TYPE "From Excel: Data"
VERSION : 0.1
   STRUCT
      kp8Stns : Array[0.."kp8StnCount"] of "From Excel: Codes Single Wip";
      hmiStns : Array[0.."hmi_station_count"] of "From Excel: Codes Multiple Wips";
   END_STRUCT;
   // hmiStns[0].wip[40].pnCode[3] := 1000;
   // hmiStns[0].wip[0].pnCode[2] := 20000;
   // hmiStns[0].wip[0].pnCode[1] := 244000;
   // hmiStns[0].wip[0].pnCode[0] := 1000;
   // hmiStns[0].pStn := 25;
   // kp8Stns[0].pStn := 0;
   // kp8Stns[0].pnCode[7] := 169000;
   // kp8Stns[2].pStn := 2;
   // kp8Stns[3].pStn := 3;
   // kp8Stns[4].pStn := 4;
   // kp8Stns[5].pStn := 5;
   // kp8Stns[7].pStn := 7;
   // kp8Stns[8].pStn := 8;
   // kp8Stns[9].pStn := 9;
   // kp8Stns[10].pStn := 10;
   // kp8Stns[11].pStn := 11;
   // kp8Stns[12].pStn := 12;
   // kp8Stns[13].pStn := 13;
   // kp8Stns[14].pStn := 14;
   // kp8Stns[15].pStn := 15;
   // kp8Stns[16].pStn := 16;
   // kp8Stns[17].pStn := 17;
   // kp8Stns[18].pStn := 18;
   // kp8Stns[19].pStn := 19;
   // kp8Stns[20].pStn := 20;
   // kp8Stns[21].pStn := 21;
   // kp8Stns[22].pStn := 22;
   // kp8Stns[23].pStn := 23;
   // kp8Stns[24].pStn := 24;
   // kp8Stns[6].pStn := 6;
   // kp8Stns[25].pStn := 30;
   // kp8Stns[26].pStn := 31;
   // kp8Stns[27].pStn := 32;
   // kp8Stns[28].pStn := 33;
   // kp8Stns[30].pStn := 35;
   // kp8Stns[31].pStn := 36;
   // kp8Stns[32].pStn := 37;
   // kp8Stns[29].pStn := 34;
   // kp8Stns[33].pStn := 38;
   // hmiStns[0].wip[40].pnCode[2] := 1000;
   // hmiStns[0].wip[40].pnCode[1] := 1000;
   // hmiStns[0].wip[40].pnCode[0] := 1000;
   // hmiStns[0].wip[39].pnCode[7] := 1000;
   // hmiStns[0].wip[39].pnCode[6] := 1000;
   // hmiStns[0].wip[39].pnCode[5] := 1000;
   // hmiStns[0].wip[39].pnCode[4] := 1000;
   // hmiStns[0].wip[39].pnCode[3] := 1000;
   // hmiStns[0].wip[39].pnCode[2] := 1000;
   // hmiStns[0].wip[39].pnCode[1] := 1000;
   // hmiStns[0].wip[39].pnCode[0] := 1000;
   // hmiStns[0].wip[38].pnCode[7] := 1000;
   // hmiStns[0].wip[38].pnCode[6] := 1000;
   // hmiStns[0].wip[38].pnCode[5] := 1000;
   // hmiStns[0].wip[38].pnCode[4] := 1000;
   // hmiStns[0].wip[38].pnCode[3] := 1000;
   // hmiStns[0].wip[38].pnCode[2] := 1000;
   // hmiStns[0].wip[38].pnCode[1] := 1000;
   // hmiStns[0].wip[38].pnCode[0] := 1000;
   // hmiStns[0].wip[37].pnCode[7] := 1000;
   // hmiStns[0].wip[37].pnCode[6] := 1000;
   // hmiStns[0].wip[37].pnCode[5] := 1000;
   // hmiStns[0].wip[37].pnCode[4] := 1000;
   // hmiStns[0].wip[37].pnCode[3] := 1000;
   // hmiStns[0].wip[37].pnCode[2] := 1000;
   // hmiStns[0].wip[37].pnCode[1] := 1000;
   // hmiStns[0].wip[37].pnCode[0] := 1000;
   // hmiStns[0].wip[36].pnCode[7] := 1000;
   // hmiStns[0].wip[36].pnCode[6] := 1000;
   // hmiStns[0].wip[36].pnCode[5] := 1000;
   // hmiStns[0].wip[36].pnCode[4] := 1000;
   // hmiStns[0].wip[36].pnCode[3] := 1000;
   // hmiStns[0].wip[36].pnCode[2] := 1000;
   // hmiStns[0].wip[36].pnCode[1] := 1000;
   // hmiStns[0].wip[36].pnCode[0] := 1000;
   // hmiStns[0].wip[35].pnCode[7] := 1000;
   // hmiStns[0].wip[35].pnCode[6] := 1000;
   // hmiStns[0].wip[35].pnCode[5] := 1000;
   // hmiStns[0].wip[35].pnCode[4] := 1000;
   // hmiStns[0].wip[35].pnCode[3] := 1000;
   // hmiStns[0].wip[35].pnCode[2] := 1000;
   // hmiStns[0].wip[35].pnCode[1] := 1000;
   // hmiStns[0].wip[35].pnCode[0] := 1000;
   // hmiStns[0].wip[34].pnCode[7] := 1000;
   // hmiStns[0].wip[34].pnCode[6] := 1000;
   // hmiStns[0].wip[34].pnCode[5] := 1000;
   // hmiStns[0].wip[34].pnCode[4] := 1000;
   // hmiStns[0].wip[34].pnCode[3] := 1000;
   // hmiStns[0].wip[34].pnCode[2] := 1000;
   // hmiStns[0].wip[34].pnCode[1] := 1000;
   // hmiStns[0].wip[34].pnCode[0] := 1000;
   // hmiStns[0].wip[33].pnCode[7] := 1000;
   // hmiStns[0].wip[33].pnCode[6] := 1000;
   // hmiStns[0].wip[33].pnCode[5] := 1000;
   // hmiStns[0].wip[33].pnCode[4] := 1000;
   // hmiStns[0].wip[33].pnCode[3] := 1000;
   // hmiStns[0].wip[33].pnCode[2] := 1000;
   // hmiStns[0].wip[33].pnCode[1] := 1000;
   // hmiStns[0].wip[33].pnCode[0] := 1000;
   // hmiStns[0].wip[32].pnCode[7] := 1000;
   // hmiStns[0].wip[32].pnCode[6] := 1000;
   // hmiStns[0].wip[32].pnCode[5] := 1000;
   // hmiStns[0].wip[32].pnCode[4] := 1000;
   // hmiStns[0].wip[32].pnCode[3] := 1000;
   // hmiStns[0].wip[32].pnCode[2] := 1000;
   // hmiStns[0].wip[32].pnCode[1] := 1000;
   // hmiStns[0].wip[32].pnCode[0] := 1000;
   // hmiStns[0].wip[31].pnCode[7] := 1000;
   // hmiStns[0].wip[31].pnCode[6] := 1000;
   // hmiStns[0].wip[31].pnCode[5] := 1000;
   // hmiStns[0].wip[31].pnCode[4] := 1000;
   // hmiStns[0].wip[31].pnCode[3] := 1000;
   // hmiStns[0].wip[31].pnCode[2] := 1000;
   // hmiStns[0].wip[31].pnCode[1] := 1000;
   // hmiStns[0].wip[31].pnCode[0] := 1000;
   // hmiStns[0].wip[30].pnCode[7] := 1000;
   // hmiStns[0].wip[30].pnCode[6] := 1000;
   // hmiStns[0].wip[30].pnCode[5] := 1000;
   // hmiStns[0].wip[30].pnCode[4] := 1000;
   // hmiStns[0].wip[30].pnCode[3] := 1000;
   // hmiStns[0].wip[30].pnCode[2] := 1000;
   // hmiStns[0].wip[30].pnCode[1] := 1000;
   // hmiStns[0].wip[30].pnCode[0] := 1000;
   // hmiStns[0].wip[29].pnCode[7] := 1000;
   // hmiStns[0].wip[29].pnCode[6] := 1000;
   // hmiStns[0].wip[29].pnCode[5] := 1000;
   // hmiStns[0].wip[29].pnCode[4] := 1000;
   // hmiStns[0].wip[29].pnCode[3] := 1000;
   // hmiStns[0].wip[29].pnCode[2] := 1000;
   // hmiStns[0].wip[29].pnCode[1] := 1000;
   // hmiStns[0].wip[29].pnCode[0] := 1000;
   // hmiStns[0].wip[28].pnCode[7] := 1000;
   // hmiStns[0].wip[28].pnCode[6] := 1000;
   // hmiStns[0].wip[28].pnCode[5] := 1000;
   // hmiStns[0].wip[28].pnCode[4] := 1000;
   // hmiStns[0].wip[28].pnCode[3] := 1000;
   // hmiStns[0].wip[28].pnCode[2] := 1000;
   // hmiStns[0].wip[28].pnCode[1] := 1000;
   // hmiStns[0].wip[28].pnCode[0] := 1000;
   // hmiStns[0].wip[27].pnCode[7] := 1000;
   // hmiStns[0].wip[27].pnCode[6] := 1000;
   // hmiStns[0].wip[27].pnCode[5] := 1000;
   // hmiStns[0].wip[27].pnCode[4] := 1000;
   // hmiStns[0].wip[27].pnCode[3] := 1000;
   // hmiStns[0].wip[27].pnCode[2] := 1000;
   // hmiStns[0].wip[27].pnCode[1] := 1000;
   // hmiStns[0].wip[27].pnCode[0] := 1000;
   // hmiStns[0].wip[26].pnCode[7] := 1000;
   // hmiStns[0].wip[26].pnCode[6] := 1000;
   // hmiStns[0].wip[26].pnCode[5] := 1000;
   // hmiStns[0].wip[26].pnCode[4] := 1000;
   // hmiStns[0].wip[26].pnCode[3] := 1000;
   // hmiStns[0].wip[26].pnCode[2] := 1000;
   // hmiStns[0].wip[26].pnCode[1] := 1000;
   // hmiStns[0].wip[26].pnCode[0] := 1000;
   // hmiStns[0].wip[25].pnCode[7] := 1000;
   // hmiStns[0].wip[25].pnCode[6] := 1000;
   // hmiStns[0].wip[25].pnCode[5] := 1000;
   // hmiStns[0].wip[25].pnCode[4] := 1000;
   // hmiStns[0].wip[25].pnCode[3] := 1000;
   // hmiStns[0].wip[25].pnCode[2] := 1000;
   // hmiStns[0].wip[25].pnCode[1] := 1000;
   // hmiStns[0].wip[25].pnCode[0] := 1000;
   // hmiStns[0].wip[24].pnCode[7] := 1000;
   // hmiStns[0].wip[24].pnCode[6] := 1000;
   // hmiStns[0].wip[24].pnCode[5] := 1000;
   // hmiStns[0].wip[24].pnCode[4] := 1000;
   // hmiStns[0].wip[24].pnCode[3] := 1000;
   // hmiStns[0].wip[24].pnCode[2] := 1000;
   // hmiStns[0].wip[24].pnCode[1] := 1000;
   // hmiStns[0].wip[24].pnCode[0] := 1000;
   // hmiStns[0].wip[23].pnCode[7] := 223000;
   // hmiStns[0].wip[23].pnCode[6] := 220000;
   // hmiStns[0].wip[23].pnCode[5] := 1000;
   // hmiStns[0].wip[23].pnCode[4] := 1000;
   // hmiStns[0].wip[23].pnCode[3] := 1000;
   // hmiStns[0].wip[23].pnCode[2] := 221000;
   // hmiStns[0].wip[23].pnCode[1] := 244000;
   // hmiStns[0].wip[23].pnCode[0] := 1000;
   // hmiStns[0].wip[22].pnCode[7] := 223000;
   // hmiStns[0].wip[22].pnCode[6] := 222000;
   // hmiStns[0].wip[22].pnCode[5] := 1000;
   // hmiStns[0].wip[22].pnCode[4] := 1000;
   // hmiStns[0].wip[22].pnCode[3] := 220000;
   // hmiStns[0].wip[22].pnCode[2] := 1000;
   // hmiStns[0].wip[22].pnCode[1] := 244000;
   // hmiStns[0].wip[22].pnCode[0] := 1000;
   // hmiStns[0].wip[21].pnCode[7] := 31000;
   // hmiStns[0].wip[21].pnCode[6] := 51000;
   // hmiStns[0].wip[21].pnCode[5] := 1000;
   // hmiStns[0].wip[21].pnCode[4] := 1000;
   // hmiStns[0].wip[21].pnCode[3] := 32000;
   // hmiStns[0].wip[21].pnCode[2] := 1000;
   // hmiStns[0].wip[21].pnCode[1] := 244000;
   // hmiStns[0].wip[21].pnCode[0] := 1000;
   // hmiStns[0].wip[20].pnCode[7] := 17000;
   // hmiStns[0].wip[20].pnCode[6] := 25000;
   // hmiStns[0].wip[20].pnCode[5] := 1000;
   // hmiStns[0].wip[20].pnCode[4] := 1000;
   // hmiStns[0].wip[20].pnCode[3] := 1000;
   // hmiStns[0].wip[20].pnCode[2] := 18000;
   // hmiStns[0].wip[20].pnCode[1] := 244000;
   // hmiStns[0].wip[20].pnCode[0] := 1000;
   // hmiStns[0].wip[19].pnCode[7] := 227000;
   // hmiStns[0].wip[19].pnCode[6] := 226000;
   // hmiStns[0].wip[19].pnCode[5] := 1000;
   // hmiStns[0].wip[19].pnCode[4] := 1000;
   // hmiStns[0].wip[19].pnCode[3] := 1000;
   // hmiStns[0].wip[19].pnCode[2] := 225000;
   // hmiStns[0].wip[19].pnCode[1] := 244000;
   // hmiStns[0].wip[19].pnCode[0] := 1000;
   // hmiStns[0].wip[18].pnCode[7] := 224000;
   // hmiStns[0].wip[18].pnCode[6] := 219000;
   // hmiStns[0].wip[18].pnCode[5] := 1000;
   // hmiStns[0].wip[18].pnCode[4] := 1000;
   // hmiStns[0].wip[18].pnCode[3] := 1000;
   // hmiStns[0].wip[18].pnCode[2] := 199000;
   // hmiStns[0].wip[18].pnCode[1] := 244000;
   // hmiStns[0].wip[18].pnCode[0] := 1000;
   // hmiStns[0].wip[17].pnCode[7] := 223000;
   // hmiStns[0].wip[17].pnCode[6] := 220000;
   // hmiStns[0].wip[17].pnCode[5] := 1000;
   // hmiStns[0].wip[17].pnCode[4] := 1000;
   // hmiStns[0].wip[17].pnCode[3] := 1000;
   // hmiStns[0].wip[17].pnCode[2] := 198000;
   // hmiStns[0].wip[17].pnCode[1] := 244000;
   // hmiStns[0].wip[17].pnCode[0] := 1000;
   // hmiStns[0].wip[16].pnCode[7] := 224000;
   // hmiStns[0].wip[16].pnCode[6] := 219000;
   // hmiStns[0].wip[16].pnCode[5] := 1000;
   // hmiStns[0].wip[16].pnCode[4] := 1000;
   // hmiStns[0].wip[16].pnCode[3] := 1000;
   // hmiStns[0].wip[16].pnCode[2] := 218000;
   // hmiStns[0].wip[16].pnCode[1] := 244000;
   // hmiStns[0].wip[16].pnCode[0] := 1000;
   // hmiStns[0].wip[15].pnCode[7] := 37000;
   // hmiStns[0].wip[15].pnCode[6] := 36000;
   // hmiStns[0].wip[15].pnCode[5] := 1000;
   // hmiStns[0].wip[15].pnCode[4] := 1000;
   // hmiStns[0].wip[15].pnCode[3] := 1000;
   // hmiStns[0].wip[15].pnCode[2] := 100000;
   // hmiStns[0].wip[15].pnCode[1] := 244000;
   // hmiStns[0].wip[15].pnCode[0] := 1000;
   // hmiStns[0].wip[14].pnCode[7] := 37000;
   // hmiStns[0].wip[14].pnCode[6] := 43000;
   // hmiStns[0].wip[14].pnCode[5] := 1000;
   // hmiStns[0].wip[14].pnCode[4] := 1000;
   // hmiStns[0].wip[14].pnCode[3] := 1000;
   // hmiStns[0].wip[14].pnCode[2] := 100000;
   // hmiStns[0].wip[14].pnCode[1] := 244000;
   // hmiStns[0].wip[14].pnCode[0] := 1000;
   // hmiStns[0].wip[13].pnCode[7] := 45000;
   // hmiStns[0].wip[13].pnCode[6] := 39000;
   // hmiStns[0].wip[13].pnCode[5] := 1000;
   // hmiStns[0].wip[13].pnCode[4] := 1000;
   // hmiStns[0].wip[13].pnCode[3] := 1000;
   // hmiStns[0].wip[13].pnCode[2] := 99000;
   // hmiStns[0].wip[13].pnCode[1] := 244000;
   // hmiStns[0].wip[13].pnCode[0] := 1000;
   // hmiStns[0].wip[12].pnCode[7] := 72000;
   // hmiStns[0].wip[12].pnCode[6] := 32000;
   // hmiStns[0].wip[12].pnCode[5] := 1000;
   // hmiStns[0].wip[12].pnCode[4] := 1000;
   // hmiStns[0].wip[12].pnCode[3] := 1000;
   // hmiStns[0].wip[12].pnCode[2] := 85000;
   // hmiStns[0].wip[12].pnCode[1] := 244000;
   // hmiStns[0].wip[12].pnCode[0] := 1000;
   // hmiStns[0].wip[11].pnCode[7] := 19000;
   // hmiStns[0].wip[11].pnCode[6] := 26000;
   // hmiStns[0].wip[11].pnCode[5] := 1000;
   // hmiStns[0].wip[11].pnCode[4] := 1000;
   // hmiStns[0].wip[11].pnCode[3] := 1000;
   // hmiStns[0].wip[11].pnCode[2] := 58000;
   // hmiStns[0].wip[11].pnCode[1] := 244000;
   // hmiStns[0].wip[11].pnCode[0] := 1000;
   // hmiStns[0].wip[10].pnCode[7] := 72000;
   // hmiStns[0].wip[10].pnCode[6] := 32000;
   // hmiStns[0].wip[10].pnCode[5] := 1000;
   // hmiStns[0].wip[10].pnCode[4] := 1000;
   // hmiStns[0].wip[10].pnCode[3] := 1000;
   // hmiStns[0].wip[10].pnCode[2] := 54000;
   // hmiStns[0].wip[10].pnCode[1] := 244000;
   // hmiStns[0].wip[10].pnCode[0] := 1000;
   // hmiStns[0].wip[9].pnCode[7] := 74000;
   // hmiStns[0].wip[9].pnCode[6] := 32000;
   // hmiStns[0].wip[9].pnCode[5] := 1000;
   // hmiStns[0].wip[9].pnCode[4] := 1000;
   // hmiStns[0].wip[9].pnCode[3] := 1000;
   // hmiStns[0].wip[9].pnCode[2] := 53000;
   // hmiStns[0].wip[9].pnCode[1] := 244000;
   // hmiStns[0].wip[9].pnCode[0] := 1000;
   // hmiStns[0].wip[8].pnCode[7] := 19000;
   // hmiStns[0].wip[8].pnCode[6] := 26000;
   // hmiStns[0].wip[8].pnCode[5] := 1000;
   // hmiStns[0].wip[8].pnCode[4] := 1000;
   // hmiStns[0].wip[8].pnCode[3] := 1000;
   // hmiStns[0].wip[8].pnCode[2] := 52000;
   // hmiStns[0].wip[8].pnCode[1] := 244000;
   // hmiStns[0].wip[8].pnCode[0] := 1000;
   // hmiStns[0].wip[7].pnCode[7] := 45000;
   // hmiStns[0].wip[7].pnCode[6] := 39000;
   // hmiStns[0].wip[7].pnCode[5] := 1000;
   // hmiStns[0].wip[7].pnCode[4] := 1000;
   // hmiStns[0].wip[7].pnCode[3] := 1000;
   // hmiStns[0].wip[7].pnCode[2] := 44000;
   // hmiStns[0].wip[7].pnCode[1] := 244000;
   // hmiStns[0].wip[7].pnCode[0] := 1000;
   // hmiStns[0].wip[6].pnCode[7] := 37000;
   // hmiStns[0].wip[6].pnCode[6] := 43000;
   // hmiStns[0].wip[6].pnCode[5] := 1000;
   // hmiStns[0].wip[6].pnCode[4] := 1000;
   // hmiStns[0].wip[6].pnCode[3] := 1000;
   // hmiStns[0].wip[6].pnCode[2] := 46000;
   // hmiStns[0].wip[6].pnCode[1] := 244000;
   // hmiStns[0].wip[6].pnCode[0] := 1000;
   // hmiStns[0].wip[5].pnCode[7] := 37000;
   // hmiStns[0].wip[5].pnCode[6] := 43000;
   // hmiStns[0].wip[5].pnCode[5] := 1000;
   // hmiStns[0].wip[5].pnCode[4] := 1000;
   // hmiStns[0].wip[5].pnCode[3] := 1000;
   // hmiStns[0].wip[5].pnCode[2] := 38000;
   // hmiStns[0].wip[5].pnCode[1] := 244000;
   // hmiStns[0].wip[5].pnCode[0] := 1000;
   // hmiStns[0].wip[4].pnCode[7] := 37000;
   // hmiStns[0].wip[4].pnCode[6] := 36000;
   // hmiStns[0].wip[4].pnCode[5] := 1000;
   // hmiStns[0].wip[4].pnCode[4] := 1000;
   // hmiStns[0].wip[4].pnCode[3] := 1000;
   // hmiStns[0].wip[4].pnCode[2] := 46000;
   // hmiStns[0].wip[4].pnCode[1] := 244000;
   // hmiStns[0].wip[4].pnCode[0] := 1000;
   // hmiStns[0].wip[3].pnCode[7] := 33000;
   // hmiStns[0].wip[3].pnCode[6] := 42000;
   // hmiStns[0].wip[3].pnCode[5] := 15000;
   // hmiStns[0].wip[3].pnCode[4] := 1000;
   // hmiStns[0].wip[3].pnCode[3] := 14000;
   // hmiStns[0].wip[3].pnCode[2] := 48000;
   // hmiStns[0].wip[3].pnCode[1] := 244000;
   // hmiStns[0].wip[3].pnCode[0] := 1000;
   // hmiStns[0].wip[2].pnCode[7] := 40000;
   // hmiStns[0].wip[2].pnCode[6] := 39000;
   // hmiStns[0].wip[2].pnCode[5] := 1000;
   // hmiStns[0].wip[2].pnCode[4] := 1000;
   // hmiStns[0].wip[2].pnCode[3] := 1000;
   // hmiStns[0].wip[2].pnCode[2] := 41000;
   // hmiStns[0].wip[2].pnCode[1] := 244000;
   // hmiStns[0].wip[2].pnCode[0] := 1000;
   // hmiStns[0].wip[1].pnCode[7] := 37000;
   // hmiStns[0].wip[1].pnCode[6] := 36000;
   // hmiStns[0].wip[1].pnCode[5] := 1000;
   // hmiStns[0].wip[1].pnCode[4] := 1000;
   // hmiStns[0].wip[1].pnCode[3] := 1000;
   // hmiStns[0].wip[1].pnCode[2] := 38000;
   // hmiStns[0].wip[1].pnCode[1] := 244000;
   // hmiStns[0].wip[1].pnCode[0] := 1000;
   // hmiStns[0].wip[0].pnCode[7] := 19000;
   // hmiStns[0].wip[0].pnCode[6] := 26000;
   // hmiStns[0].wip[0].pnCode[5] := 1000;
   // hmiStns[0].wip[0].pnCode[4] := 1000;
   // hmiStns[0].wip[0].pnCode[3] := 1000;
   // kp8Stns[1].pnCode[0] := 1000;
   // kp8Stns[0].pnCode[1] := 1000;
   // kp8Stns[0].pnCode[0] := 1000;
   // kp8Stns[0].pnCode[2] := 1000;
   // kp8Stns[0].pnCode[3] := 173000;
   // kp8Stns[0].pnCode[4] := 1000;
   // kp8Stns[0].pnCode[5] := 1000;
   // kp8Stns[0].pnCode[6] := 1000;
   // kp8Stns[1].pnCode[1] := 1000;
   // kp8Stns[1].pnCode[2] := 184000;
   // kp8Stns[1].pnCode[3] := 210000;
   // kp8Stns[1].pnCode[4] := 1000;
   // kp8Stns[1].pnCode[5] := 1000;
   // kp8Stns[1].pnCode[6] := 181000;
   // kp8Stns[1].pnCode[7] := 167000;
   // kp8Stns[1].pStn := 1;
   // kp8Stns[2].pnCode[0] := 1000;
   // kp8Stns[2].pnCode[1] := 183000;
   // kp8Stns[2].pnCode[2] := 182000;
   // kp8Stns[2].pnCode[3] := 216000;
   // kp8Stns[2].pnCode[4] := 1000;
   // kp8Stns[2].pnCode[5] := 185000;
   // kp8Stns[2].pnCode[6] := 217000;
   // kp8Stns[2].pnCode[7] := 215000;
   // kp8Stns[3].pnCode[0] := 1000;
   // kp8Stns[3].pnCode[1] := 193000;
   // kp8Stns[3].pnCode[2] := 192000;
   // kp8Stns[3].pnCode[3] := 189000;
   // kp8Stns[3].pnCode[4] := 1000;
   // kp8Stns[3].pnCode[5] := 191000;
   // kp8Stns[3].pnCode[6] := 188000;
   // kp8Stns[3].pnCode[7] := 190000;
   // kp8Stns[4].pnCode[0] := 1000;
   // kp8Stns[4].pnCode[1] := 1000;
   // kp8Stns[4].pnCode[2] := 1000;
   // kp8Stns[4].pnCode[3] := 1000;
   // kp8Stns[4].pnCode[4] := 1000;
   // kp8Stns[4].pnCode[5] := 1000;
   // kp8Stns[4].pnCode[6] := 1000;
   // kp8Stns[4].pnCode[7] := 195000;
   // kp8Stns[5].pnCode[0] := 1000;
   // kp8Stns[5].pnCode[1] := 194000;
   // kp8Stns[5].pnCode[2] := 196000;
   // kp8Stns[5].pnCode[3] := 177000;
   // kp8Stns[5].pnCode[4] := 1000;
   // kp8Stns[5].pnCode[5] := 197000;
   // kp8Stns[5].pnCode[6] := 178000;
   // kp8Stns[5].pnCode[7] := 176000;
   // kp8Stns[6].pnCode[0] := 1000;
   // kp8Stns[6].pnCode[1] := 209000;
   // kp8Stns[6].pnCode[2] := 208000;
   // kp8Stns[6].pnCode[3] := 211000;
   // kp8Stns[6].pnCode[4] := 1000;
   // kp8Stns[6].pnCode[5] := 212000;
   // kp8Stns[6].pnCode[6] := 207000;
   // kp8Stns[6].pnCode[7] := 206000;
   // kp8Stns[7].pnCode[0] := 1000;
   // kp8Stns[7].pnCode[1] := 1000;
   // kp8Stns[7].pnCode[2] := 1000;
   // kp8Stns[7].pnCode[3] := 175000;
   // kp8Stns[7].pnCode[4] := 1000;
   // kp8Stns[7].pnCode[5] := 1000;
   // kp8Stns[7].pnCode[6] := 168000;
   // kp8Stns[7].pnCode[7] := 170000;
   // kp8Stns[8].pnCode[0] := 1000;
   // kp8Stns[8].pnCode[1] := 1000;
   // kp8Stns[8].pnCode[2] := 1000;
   // kp8Stns[8].pnCode[3] := 205000;
   // kp8Stns[8].pnCode[4] := 1000;
   // kp8Stns[8].pnCode[5] := 1000;
   // kp8Stns[8].pnCode[6] := 174000;
   // kp8Stns[8].pnCode[7] := 187000;
   // kp8Stns[9].pnCode[0] := 1000;
   // kp8Stns[9].pnCode[1] := 1000;
   // kp8Stns[9].pnCode[2] := 1000;
   // kp8Stns[9].pnCode[3] := 214000;
   // kp8Stns[9].pnCode[4] := 1000;
   // kp8Stns[9].pnCode[5] := 1000;
   // kp8Stns[9].pnCode[6] := 1000;
   // kp8Stns[9].pnCode[7] := 213000;
   // kp8Stns[10].pnCode[0] := 1000;
   // kp8Stns[10].pnCode[1] := 1000;
   // kp8Stns[10].pnCode[2] := 1000;
   // kp8Stns[10].pnCode[3] := 171000;
   // kp8Stns[10].pnCode[4] := 1000;
   // kp8Stns[10].pnCode[5] := 1000;
   // kp8Stns[10].pnCode[6] := 243000;
   // kp8Stns[10].pnCode[7] := 172000;
   // kp8Stns[11].pnCode[0] := 1000;
   // kp8Stns[11].pnCode[1] := 1000;
   // kp8Stns[11].pnCode[2] := 1000;
   // kp8Stns[11].pnCode[3] := 78000;
   // kp8Stns[11].pnCode[4] := 1000;
   // kp8Stns[11].pnCode[5] := 1000;
   // kp8Stns[11].pnCode[6] := 66000;
   // kp8Stns[11].pnCode[7] := 21000;
   // kp8Stns[12].pnCode[0] := 1000;
   // kp8Stns[12].pnCode[1] := 81000;
   // kp8Stns[12].pnCode[2] := 87000;
   // kp8Stns[12].pnCode[3] := 60000;
   // kp8Stns[12].pnCode[4] := 1000;
   // kp8Stns[12].pnCode[5] := 80000;
   // kp8Stns[12].pnCode[6] := 56000;
   // kp8Stns[12].pnCode[7] := 55000;
   // kp8Stns[13].pnCode[0] := 1000;
   // kp8Stns[13].pnCode[1] := 1000;
   // kp8Stns[13].pnCode[2] := 70000;
   // kp8Stns[13].pnCode[3] := 90000;
   // kp8Stns[13].pnCode[4] := 1000;
   // kp8Stns[13].pnCode[5] := 1000;
   // kp8Stns[13].pnCode[6] := 91000;
   // kp8Stns[13].pnCode[7] := 89000;
   // kp8Stns[14].pnCode[0] := 1000;
   // kp8Stns[14].pnCode[1] := 1000;
   // kp8Stns[14].pnCode[2] := 65000;
   // kp8Stns[14].pnCode[3] := 88000;
   // kp8Stns[14].pnCode[4] := 1000;
   // kp8Stns[14].pnCode[5] := 64000;
   // kp8Stns[14].pnCode[6] := 83000;
   // kp8Stns[14].pnCode[7] := 63000;
   // kp8Stns[15].pnCode[0] := 1000;
   // kp8Stns[15].pnCode[1] := 50000;
   // kp8Stns[15].pnCode[2] := 77000;
   // kp8Stns[15].pnCode[3] := 29000;
   // kp8Stns[15].pnCode[4] := 1000;
   // kp8Stns[15].pnCode[5] := 82000;
   // kp8Stns[15].pnCode[6] := 69000;
   // kp8Stns[15].pnCode[7] := 75000;
   // kp8Stns[16].pnCode[0] := 1000;
   // kp8Stns[16].pnCode[1] := 1000;
   // kp8Stns[16].pnCode[2] := 1000;
   // kp8Stns[16].pnCode[3] := 92000;
   // kp8Stns[16].pnCode[4] := 1000;
   // kp8Stns[16].pnCode[5] := 1000;
   // kp8Stns[16].pnCode[6] := 94000;
   // kp8Stns[16].pnCode[7] := 95068;
   // kp8Stns[17].pnCode[0] := 1000;
   // kp8Stns[17].pnCode[1] := 1000;
   // kp8Stns[17].pnCode[2] := 84000;
   // kp8Stns[17].pnCode[3] := 35000;
   // kp8Stns[17].pnCode[4] := 1000;
   // kp8Stns[17].pnCode[5] := 1000;
   // kp8Stns[17].pnCode[6] := 76000;
   // kp8Stns[17].pnCode[7] := 30000;
   // kp8Stns[18].pnCode[0] := 1000;
   // kp8Stns[18].pnCode[1] := 1000;
   // kp8Stns[18].pnCode[2] := 1000;
   // kp8Stns[18].pnCode[3] := 188135;
   // kp8Stns[18].pnCode[4] := 1000;
   // kp8Stns[18].pnCode[5] := 1000;
   // kp8Stns[18].pnCode[6] := 285162;
   // kp8Stns[18].pnCode[7] := 96000;
   // kp8Stns[19].pnCode[0] := 1000;
   // kp8Stns[19].pnCode[1] := 79000;
   // kp8Stns[19].pnCode[2] := 86000;
   // kp8Stns[19].pnCode[3] := 22000;
   // kp8Stns[19].pnCode[4] := 1000;
   // kp8Stns[19].pnCode[5] := 98000;
   // kp8Stns[19].pnCode[6] := 61000;
   // kp8Stns[19].pnCode[7] := 49000;
   // kp8Stns[20].pnCode[0] := 1000;
   // kp8Stns[20].pnCode[1] := 1000;
   // kp8Stns[20].pnCode[2] := 1000;
   // kp8Stns[20].pnCode[3] := 1000;
   // kp8Stns[20].pnCode[4] := 1000;
   // kp8Stns[20].pnCode[5] := 1000;
   // kp8Stns[20].pnCode[6] := 1000;
   // kp8Stns[20].pnCode[7] := 245000;
   // kp8Stns[21].pnCode[0] := 1000;
   // kp8Stns[21].pnCode[1] := 1000;
   // kp8Stns[21].pnCode[2] := 1000;
   // kp8Stns[21].pnCode[3] := 246000;
   // kp8Stns[21].pnCode[4] := 1000;
   // kp8Stns[21].pnCode[5] := 1000;
   // kp8Stns[21].pnCode[6] := 1000;
   // kp8Stns[21].pnCode[7] := 12000;
   // kp8Stns[22].pnCode[0] := 1000;
   // kp8Stns[22].pnCode[1] := 1000;
   // kp8Stns[22].pnCode[2] := 1000;
   // kp8Stns[22].pnCode[3] := 23000;
   // kp8Stns[22].pnCode[4] := 1000;
   // kp8Stns[22].pnCode[5] := 1000;
   // kp8Stns[22].pnCode[6] := 47000;
   // kp8Stns[22].pnCode[7] := 62000;
   // kp8Stns[23].pnCode[0] := 1000;
   // kp8Stns[23].pnCode[1] := 1000;
   // kp8Stns[23].pnCode[2] := 1000;
   // kp8Stns[23].pnCode[3] := 1000;
   // kp8Stns[23].pnCode[4] := 1000;
   // kp8Stns[23].pnCode[5] := 1000;
   // kp8Stns[23].pnCode[6] := 1000;
   // kp8Stns[23].pnCode[7] := 13000;
   // kp8Stns[24].pnCode[0] := 1000;
   // kp8Stns[24].pnCode[1] := 1000;
   // kp8Stns[24].pnCode[2] := 1000;
   // kp8Stns[24].pnCode[3] := 1000;
   // kp8Stns[24].pnCode[4] := 1000;
   // kp8Stns[24].pnCode[5] := 1000;
   // kp8Stns[24].pnCode[6] := 1000;
   // kp8Stns[24].pnCode[7] := 28000;
   // kp8Stns[25].pnCode[0] := 1000;
   // kp8Stns[25].pnCode[1] := 1000;
   // kp8Stns[25].pnCode[2] := 1000;
   // kp8Stns[25].pnCode[3] := 1000;
   // kp8Stns[25].pnCode[4] := 1000;
   // kp8Stns[25].pnCode[5] := 1000;
   // kp8Stns[25].pnCode[6] := 1000;
   // kp8Stns[25].pnCode[7] := 57000;
   // hmiStns[0].wip[40].pnCode[4] := 1000;
   // hmiStns[0].wip[40].pnCode[5] := 1000;
   // hmiStns[0].wip[40].pnCode[6] := 1000;
   // hmiStns[0].wip[40].pnCode[7] := 1000;
   // hmiStns[0].wip[41].pnCode[0] := 1000;
   // hmiStns[0].wip[41].pnCode[1] := 1000;
   // hmiStns[0].wip[41].pnCode[2] := 1000;
   // hmiStns[0].wip[41].pnCode[3] := 1000;
   // hmiStns[0].wip[41].pnCode[4] := 1000;
   // hmiStns[0].wip[41].pnCode[5] := 1000;
   // hmiStns[0].wip[41].pnCode[6] := 1000;
   // hmiStns[0].wip[41].pnCode[7] := 1000;
   // hmiStns[0].wip[42].pnCode[0] := 1000;
   // hmiStns[0].wip[42].pnCode[1] := 1000;
   // hmiStns[0].wip[42].pnCode[2] := 1000;
   // hmiStns[0].wip[42].pnCode[3] := 1000;
   // hmiStns[0].wip[42].pnCode[4] := 1000;
   // hmiStns[0].wip[42].pnCode[5] := 1000;
   // hmiStns[0].wip[42].pnCode[6] := 1000;
   // hmiStns[0].wip[42].pnCode[7] := 1000;
   // hmiStns[0].wip[43].pnCode[0] := 1000;
   // hmiStns[0].wip[43].pnCode[1] := 1000;
   // hmiStns[0].wip[43].pnCode[2] := 1000;
   // hmiStns[0].wip[43].pnCode[3] := 1000;
   // hmiStns[0].wip[43].pnCode[4] := 1000;
   // hmiStns[0].wip[43].pnCode[5] := 1000;
   // hmiStns[0].wip[43].pnCode[6] := 1000;
   // hmiStns[0].wip[43].pnCode[7] := 1000;
   // hmiStns[0].wip[44].pnCode[0] := 1000;
   // hmiStns[0].wip[44].pnCode[1] := 1000;
   // hmiStns[0].wip[44].pnCode[2] := 1000;
   // hmiStns[0].wip[44].pnCode[3] := 1000;
   // hmiStns[0].wip[44].pnCode[4] := 1000;
   // hmiStns[0].wip[44].pnCode[5] := 1000;
   // hmiStns[0].wip[44].pnCode[6] := 1000;
   // hmiStns[0].wip[44].pnCode[7] := 1000;
   // hmiStns[0].wip[45].pnCode[0] := 1000;
   // hmiStns[0].wip[45].pnCode[1] := 1000;
   // hmiStns[0].wip[45].pnCode[2] := 1000;
   // hmiStns[0].wip[45].pnCode[3] := 1000;
   // hmiStns[0].wip[45].pnCode[4] := 1000;
   // hmiStns[0].wip[45].pnCode[5] := 1000;
   // hmiStns[0].wip[45].pnCode[6] := 1000;
   // hmiStns[0].wip[45].pnCode[7] := 1000;
   // hmiStns[0].wip[46].pnCode[0] := 1000;
   // hmiStns[0].wip[46].pnCode[1] := 1000;
   // hmiStns[0].wip[46].pnCode[2] := 1000;
   // hmiStns[0].wip[46].pnCode[3] := 1000;
   // hmiStns[0].wip[46].pnCode[4] := 1000;
   // hmiStns[0].wip[46].pnCode[5] := 1000;
   // hmiStns[0].wip[46].pnCode[6] := 1000;
   // hmiStns[0].wip[46].pnCode[7] := 1000;
   // hmiStns[0].wip[47].pnCode[0] := 1000;
   // hmiStns[0].wip[47].pnCode[1] := 1000;
   // hmiStns[0].wip[47].pnCode[2] := 1000;
   // hmiStns[0].wip[47].pnCode[3] := 1000;
   // hmiStns[0].wip[47].pnCode[4] := 1000;
   // hmiStns[0].wip[47].pnCode[5] := 1000;
   // hmiStns[0].wip[47].pnCode[6] := 1000;
   // hmiStns[0].wip[47].pnCode[7] := 1000;
   // hmiStns[0].wip[48].pnCode[0] := 1000;
   // hmiStns[0].wip[48].pnCode[1] := 1000;
   // hmiStns[0].wip[48].pnCode[2] := 1000;
   // hmiStns[0].wip[48].pnCode[3] := 1000;
   // hmiStns[0].wip[48].pnCode[4] := 1000;
   // hmiStns[0].wip[48].pnCode[5] := 1000;
   // hmiStns[0].wip[48].pnCode[6] := 1000;
   // hmiStns[0].wip[48].pnCode[7] := 1000;
   // hmiStns[0].wip[49].pnCode[0] := 1000;
   // hmiStns[0].wip[49].pnCode[1] := 1000;
   // hmiStns[0].wip[49].pnCode[2] := 1000;
   // hmiStns[0].wip[49].pnCode[3] := 1000;
   // hmiStns[0].wip[49].pnCode[4] := 1000;
   // hmiStns[0].wip[49].pnCode[5] := 1000;
   // hmiStns[0].wip[49].pnCode[6] := 1000;
   // hmiStns[0].wip[49].pnCode[7] := 1000;
   // hmiStns[1].pStn := 26;
   // hmiStns[1].wip[0].pnCode[0] := 1000;
   // hmiStns[1].wip[0].pnCode[1] := 244000;
   // hmiStns[1].wip[0].pnCode[2] := 46000;
   // hmiStns[1].wip[0].pnCode[3] := 1000;
   // hmiStns[1].wip[0].pnCode[4] := 1000;
   // hmiStns[1].wip[0].pnCode[5] := 1000;
   // hmiStns[1].wip[0].pnCode[6] := 43000;
   // hmiStns[1].wip[0].pnCode[7] := 37000;
   // hmiStns[1].wip[1].pnCode[0] := 1000;
   // hmiStns[1].wip[1].pnCode[1] := 244000;
   // hmiStns[1].wip[1].pnCode[2] := 100000;
   // hmiStns[1].wip[1].pnCode[3] := 1000;
   // hmiStns[1].wip[1].pnCode[4] := 1000;
   // hmiStns[1].wip[1].pnCode[5] := 1000;
   // hmiStns[1].wip[1].pnCode[6] := 43000;
   // hmiStns[1].wip[1].pnCode[7] := 37000;
   // hmiStns[1].wip[2].pnCode[0] := 1000;
   // hmiStns[1].wip[2].pnCode[1] := 244000;
   // hmiStns[1].wip[2].pnCode[2] := 100000;
   // hmiStns[1].wip[2].pnCode[3] := 1000;
   // hmiStns[1].wip[2].pnCode[4] := 1000;
   // hmiStns[1].wip[2].pnCode[5] := 1000;
   // hmiStns[1].wip[2].pnCode[6] := 36000;
   // hmiStns[1].wip[2].pnCode[7] := 37000;
   // hmiStns[1].wip[3].pnCode[0] := 1000;
   // hmiStns[1].wip[3].pnCode[1] := 244000;
   // hmiStns[1].wip[3].pnCode[2] := 15000;
   // hmiStns[1].wip[3].pnCode[3] := 1000;
   // hmiStns[1].wip[3].pnCode[4] := 1000;
   // hmiStns[1].wip[3].pnCode[5] := 16000;
   // hmiStns[1].wip[3].pnCode[6] := 24000;
   // hmiStns[1].wip[3].pnCode[7] := 14000;
   // hmiStns[1].wip[4].pnCode[0] := 1000;
   // hmiStns[1].wip[4].pnCode[1] := 244000;
   // hmiStns[1].wip[4].pnCode[2] := 15000;
   // hmiStns[1].wip[4].pnCode[3] := 14000;
   // hmiStns[1].wip[4].pnCode[4] := 1000;
   // hmiStns[1].wip[4].pnCode[5] := 48000;
   // hmiStns[1].wip[4].pnCode[6] := 34000;
   // hmiStns[1].wip[4].pnCode[7] := 33000;
   // hmiStns[1].wip[5].pnCode[0] := 1000;
   // hmiStns[1].wip[5].pnCode[1] := 244000;
   // hmiStns[1].wip[5].pnCode[2] := 15000;
   // hmiStns[1].wip[5].pnCode[3] := 1000;
   // hmiStns[1].wip[5].pnCode[4] := 1000;
   // hmiStns[1].wip[5].pnCode[5] := 16000;
   // hmiStns[1].wip[5].pnCode[6] := 34000;
   // hmiStns[1].wip[5].pnCode[7] := 14000;
   // hmiStns[1].wip[6].pnCode[0] := 1000;
   // hmiStns[1].wip[6].pnCode[1] := 244000;
   // hmiStns[1].wip[6].pnCode[2] := 71000;
   // hmiStns[1].wip[6].pnCode[3] := 74000;
   // hmiStns[1].wip[6].pnCode[4] := 1000;
   // hmiStns[1].wip[6].pnCode[5] := 59000;
   // hmiStns[1].wip[6].pnCode[6] := 42000;
   // hmiStns[1].wip[6].pnCode[7] := 73000;
   // hmiStns[1].wip[7].pnCode[0] := 1000;
   // hmiStns[1].wip[7].pnCode[1] := 244000;
   // hmiStns[1].wip[7].pnCode[2] := 229000;
   // hmiStns[1].wip[7].pnCode[3] := 232000;
   // hmiStns[1].wip[7].pnCode[4] := 1000;
   // hmiStns[1].wip[7].pnCode[5] := 230000;
   // hmiStns[1].wip[7].pnCode[6] := 228000;
   // hmiStns[1].wip[7].pnCode[7] := 231000;
   // hmiStns[1].wip[8].pnCode[0] := 1000;
   // hmiStns[1].wip[8].pnCode[1] := 244000;
   // hmiStns[1].wip[8].pnCode[2] := 234000;
   // hmiStns[1].wip[8].pnCode[3] := 1000;
   // hmiStns[1].wip[8].pnCode[4] := 1000;
   // hmiStns[1].wip[8].pnCode[5] := 230000;
   // hmiStns[1].wip[8].pnCode[6] := 233000;
   // hmiStns[1].wip[8].pnCode[7] := 232000;
   // hmiStns[1].wip[9].pnCode[0] := 1000;
   // hmiStns[1].wip[9].pnCode[1] := 244000;
   // hmiStns[1].wip[9].pnCode[2] := 237000;
   // hmiStns[1].wip[9].pnCode[3] := 1000;
   // hmiStns[1].wip[9].pnCode[4] := 1000;
   // hmiStns[1].wip[9].pnCode[5] := 238000;
   // hmiStns[1].wip[9].pnCode[6] := 235000;
   // hmiStns[1].wip[9].pnCode[7] := 236000;
   // hmiStns[1].wip[10].pnCode[0] := 1000;
   // hmiStns[1].wip[10].pnCode[1] := 244000;
   // hmiStns[1].wip[10].pnCode[2] := 165000;
   // hmiStns[1].wip[10].pnCode[3] := 1000;
   // hmiStns[1].wip[10].pnCode[4] := 1000;
   // hmiStns[1].wip[10].pnCode[5] := 166000;
   // hmiStns[1].wip[10].pnCode[6] := 235000;
   // hmiStns[1].wip[10].pnCode[7] := 236000;
   // hmiStns[1].wip[11].pnCode[0] := 1000;
   // hmiStns[1].wip[11].pnCode[1] := 244000;
   // hmiStns[1].wip[11].pnCode[2] := 202000;
   // hmiStns[1].wip[11].pnCode[3] := 1000;
   // hmiStns[1].wip[11].pnCode[4] := 1000;
   // hmiStns[1].wip[11].pnCode[5] := 201000;
   // hmiStns[1].wip[11].pnCode[6] := 235000;
   // hmiStns[1].wip[11].pnCode[7] := 236000;
   // hmiStns[1].wip[12].pnCode[0] := 1000;
   // hmiStns[1].wip[12].pnCode[1] := 244000;
   // hmiStns[1].wip[12].pnCode[2] := 241000;
   // hmiStns[1].wip[12].pnCode[3] := 1000;
   // hmiStns[1].wip[12].pnCode[4] := 1000;
   // hmiStns[1].wip[12].pnCode[5] := 242000;
   // hmiStns[1].wip[12].pnCode[6] := 239000;
   // hmiStns[1].wip[12].pnCode[7] := 240000;
   // hmiStns[1].wip[13].pnCode[0] := 1000;
   // hmiStns[1].wip[13].pnCode[1] := 244000;
   // hmiStns[1].wip[13].pnCode[2] := 71000;
   // hmiStns[1].wip[13].pnCode[3] := 73000;
   // hmiStns[1].wip[13].pnCode[4] := 1000;
   // hmiStns[1].wip[13].pnCode[5] := 59000;
   // hmiStns[1].wip[13].pnCode[6] := 34000;
   // hmiStns[1].wip[13].pnCode[7] := 74000;
   // hmiStns[1].wip[14].pnCode[0] := 1000;
   // hmiStns[1].wip[14].pnCode[1] := 1000;
   // hmiStns[1].wip[14].pnCode[2] := 1000;
   // hmiStns[1].wip[14].pnCode[3] := 1000;
   // hmiStns[1].wip[14].pnCode[4] := 1000;
   // hmiStns[1].wip[14].pnCode[5] := 1000;
   // hmiStns[1].wip[14].pnCode[6] := 1000;
   // hmiStns[1].wip[14].pnCode[7] := 1000;
   // hmiStns[1].wip[15].pnCode[0] := 1000;
   // hmiStns[1].wip[15].pnCode[1] := 1000;
   // hmiStns[1].wip[15].pnCode[2] := 1000;
   // hmiStns[1].wip[15].pnCode[3] := 1000;
   // hmiStns[1].wip[15].pnCode[4] := 1000;
   // hmiStns[1].wip[15].pnCode[5] := 1000;
   // hmiStns[1].wip[15].pnCode[6] := 1000;
   // hmiStns[1].wip[15].pnCode[7] := 1000;
   // hmiStns[1].wip[16].pnCode[0] := 1000;
   // hmiStns[1].wip[16].pnCode[1] := 1000;
   // hmiStns[1].wip[16].pnCode[2] := 1000;
   // hmiStns[1].wip[16].pnCode[3] := 1000;
   // hmiStns[1].wip[16].pnCode[4] := 1000;
   // hmiStns[1].wip[16].pnCode[5] := 1000;
   // hmiStns[1].wip[16].pnCode[6] := 1000;
   // hmiStns[1].wip[16].pnCode[7] := 1000;
   // hmiStns[1].wip[17].pnCode[0] := 1000;
   // hmiStns[1].wip[17].pnCode[1] := 1000;
   // hmiStns[1].wip[17].pnCode[2] := 1000;
   // hmiStns[1].wip[17].pnCode[3] := 1000;
   // hmiStns[1].wip[17].pnCode[4] := 1000;
   // hmiStns[1].wip[17].pnCode[5] := 1000;
   // hmiStns[1].wip[17].pnCode[6] := 1000;
   // hmiStns[1].wip[17].pnCode[7] := 1000;
   // hmiStns[1].wip[18].pnCode[0] := 1000;
   // hmiStns[1].wip[18].pnCode[1] := 1000;
   // hmiStns[1].wip[18].pnCode[2] := 1000;